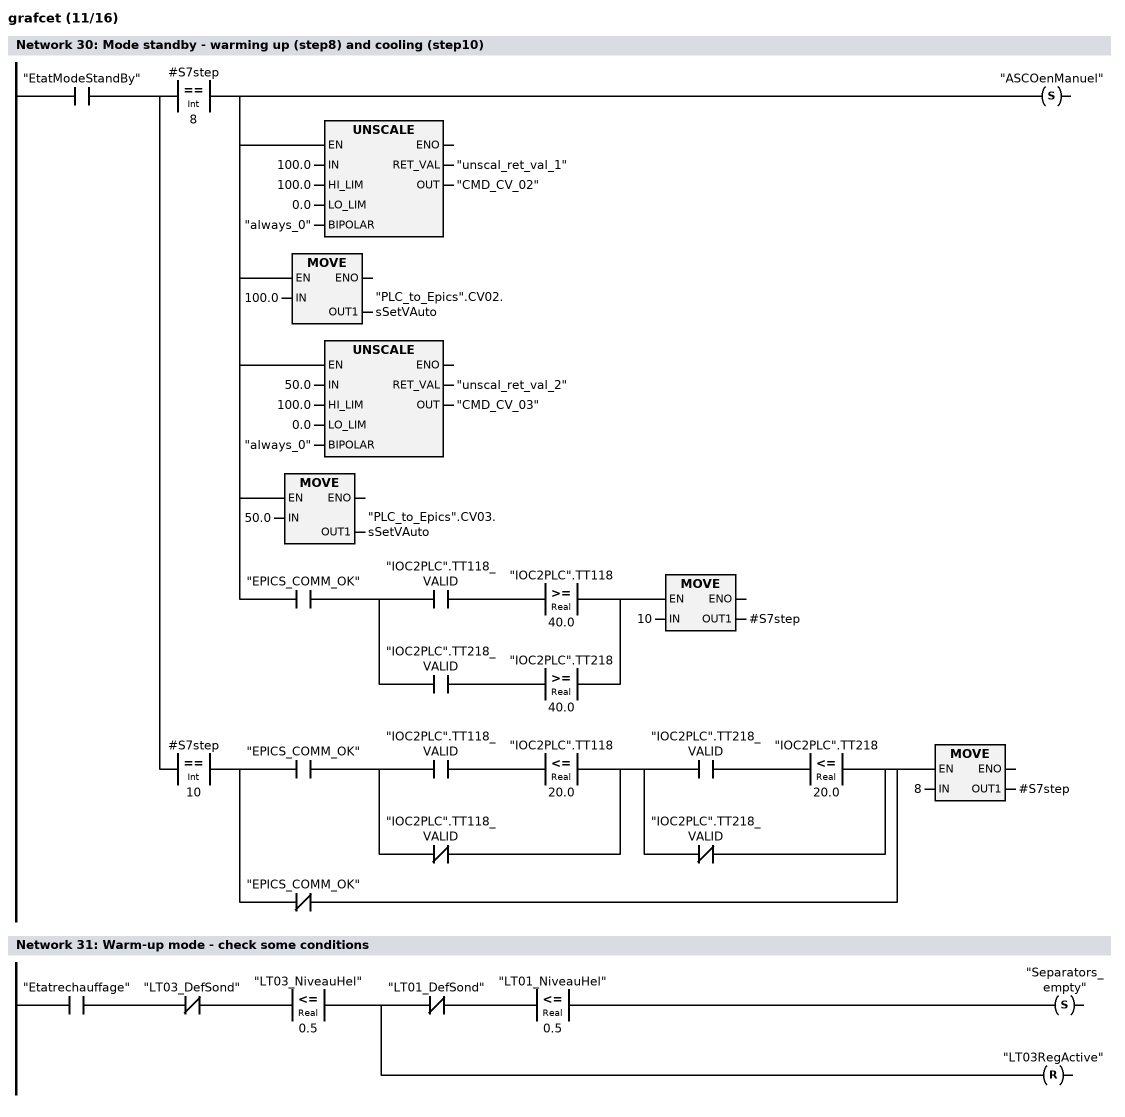
   #_w1 := "EtatModeStandBy" AND (#S7step = 8);
   IF #_w1 THEN "ASCOenManuel" := TRUE; END_IF;
   #_w2 := "EtatModeStandBy";
   IF #_w1 THEN
       "unscal_ret_val_1" := UNSCALE(IN := 100.0,
                               HI_LIM := 100.0,
                               LO_LIM := 0.0,
                               BIPOLAR := "always_0",
                               OUT => "CMD_CV_02");
       "PLC_to_Epics".CV02.sSetVAuto := 100.0;
       "unscal_ret_val_2" := UNSCALE(IN := 50.0,
                               HI_LIM := 100.0,
                               LO_LIM := 0.0,
                               BIPOLAR := "always_0",
                               OUT => "CMD_CV_03");
       "PLC_to_Epics".CV03.sSetVAuto := 50.0;
   END_IF;
   IF #_w1 AND "EPICS_COMM_OK" AND (("IOC2PLC".TT118_VALID AND ("IOC2PLC".TT118 >= 40.0)) OR ("IOC2PLC".TT218_VALID AND ("IOC2PLC".TT218 >= 40.0))) THEN
       #S7step := 10;
   END_IF;
   IF #_w2 AND (#S7step = 10) AND (("EPICS_COMM_OK" AND (("IOC2PLC".TT118_VALID AND ("IOC2PLC".TT118 <= 20.0)) OR NOT "IOC2PLC".TT118_VALID) AND (("IOC2PLC".TT218_VALID AND ("IOC2PLC".TT218 <= 20.0)) OR NOT "IOC2PLC".TT218_VALID)) OR NOT "EPICS_COMM_OK") THEN
       #S7step := 8;
   END_IF;
END_REGION

REGION Network 31: Warm-up mode - check some conditions
   #_w1 := "Etatrechauffage" AND NOT "LT03_DefSond" AND ("LT03_NiveauHel" <= 0.5);
   IF #_w1 AND NOT "LT01_DefSond" AND ("LT01_NiveauHel" <= 0.5) THEN "Separators_empty" := TRUE; END_IF;
   IF #_w1 THEN "LT03RegActive" := FALSE; END_IF;
END_REGION

REGION Network 32: Warm-up: set-up the settings of CV01-CV04
   // Set-up the settings depending on the LHe levels in the phase separators
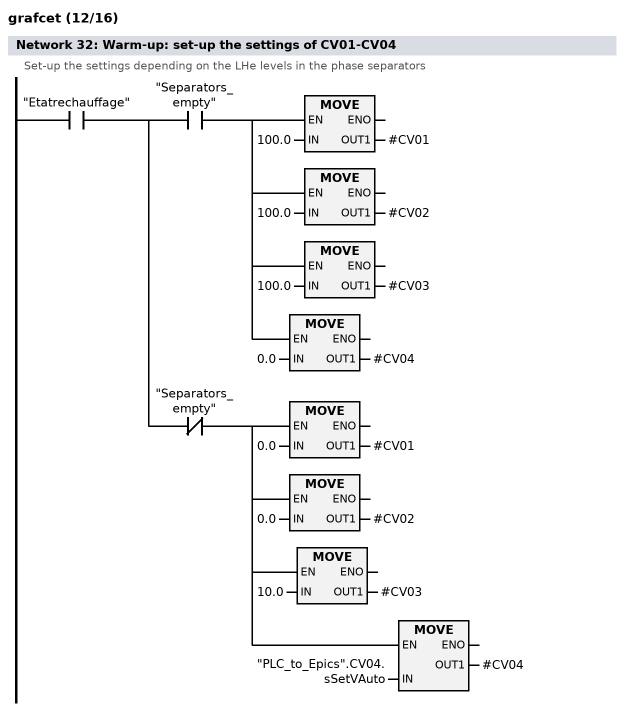
   RUNG wire#powerrail
      Contact( "Etatrechauffage" )
      wire#w1
      Contact( "Separators_empty" )
      wire#w2
      { S7_GenerateENO := "TRUE" } Move(in := 100.0, out1 => #CV01)
   END_RUNG
   RUNG wire#w2
      { S7_GenerateENO := "TRUE" } Move(in := 100.0, out1 => #CV02)
   END_RUNG
   RUNG wire#w2
      { S7_GenerateENO := "TRUE" } Move(in := 100.0, out1 => #CV03)
   END_RUNG
   RUNG wire#w2
      { S7_GenerateENO := "TRUE" } Move(in := 0.0, out1 => #CV04)
   END_RUNG
   RUNG wire#w1
      I_Contact( "Separators_empty" )
      wire#w3
      { S7_GenerateENO := "TRUE" } Move(in := 0.0, out1 => #CV01)
   END_RUNG
   RUNG wire#w3
      { S7_GenerateENO := "TRUE" } Move(in := 0.0, out1 => #CV02)
   END_RUNG
   RUNG wire#w3
      { S7_GenerateENO := "TRUE" } Move(in := 10.0, out1 => #CV03)
   END_RUNG
   RUNG wire#w3
      { S7_GenerateENO := "TRUE" } Move(in := "PLC_to_Epics".CV04.sSetVAuto, out1 => #CV04)
   END_RUNG
   // the same network as SCL:
   IF "Etatrechauffage" AND "Separators_empty" THEN
       #CV01 := 100.0;
       #CV02 := 100.0;
       #CV03 := 100.0;
       #CV04 := 0.0;
   END_IF;
   IF "Etatrechauffage" AND NOT "Separators_empty" THEN
       #CV01 := 0.0;
       #CV02 := 0.0;
       #CV03 := 10.0;
       #CV04 := "PLC_to_Epics".CV04.sSetVAuto;
   END_IF;
END_REGION

REGION Network 33: Mode Rechauffage
   // The heaters are handled in Manage_HEATERS
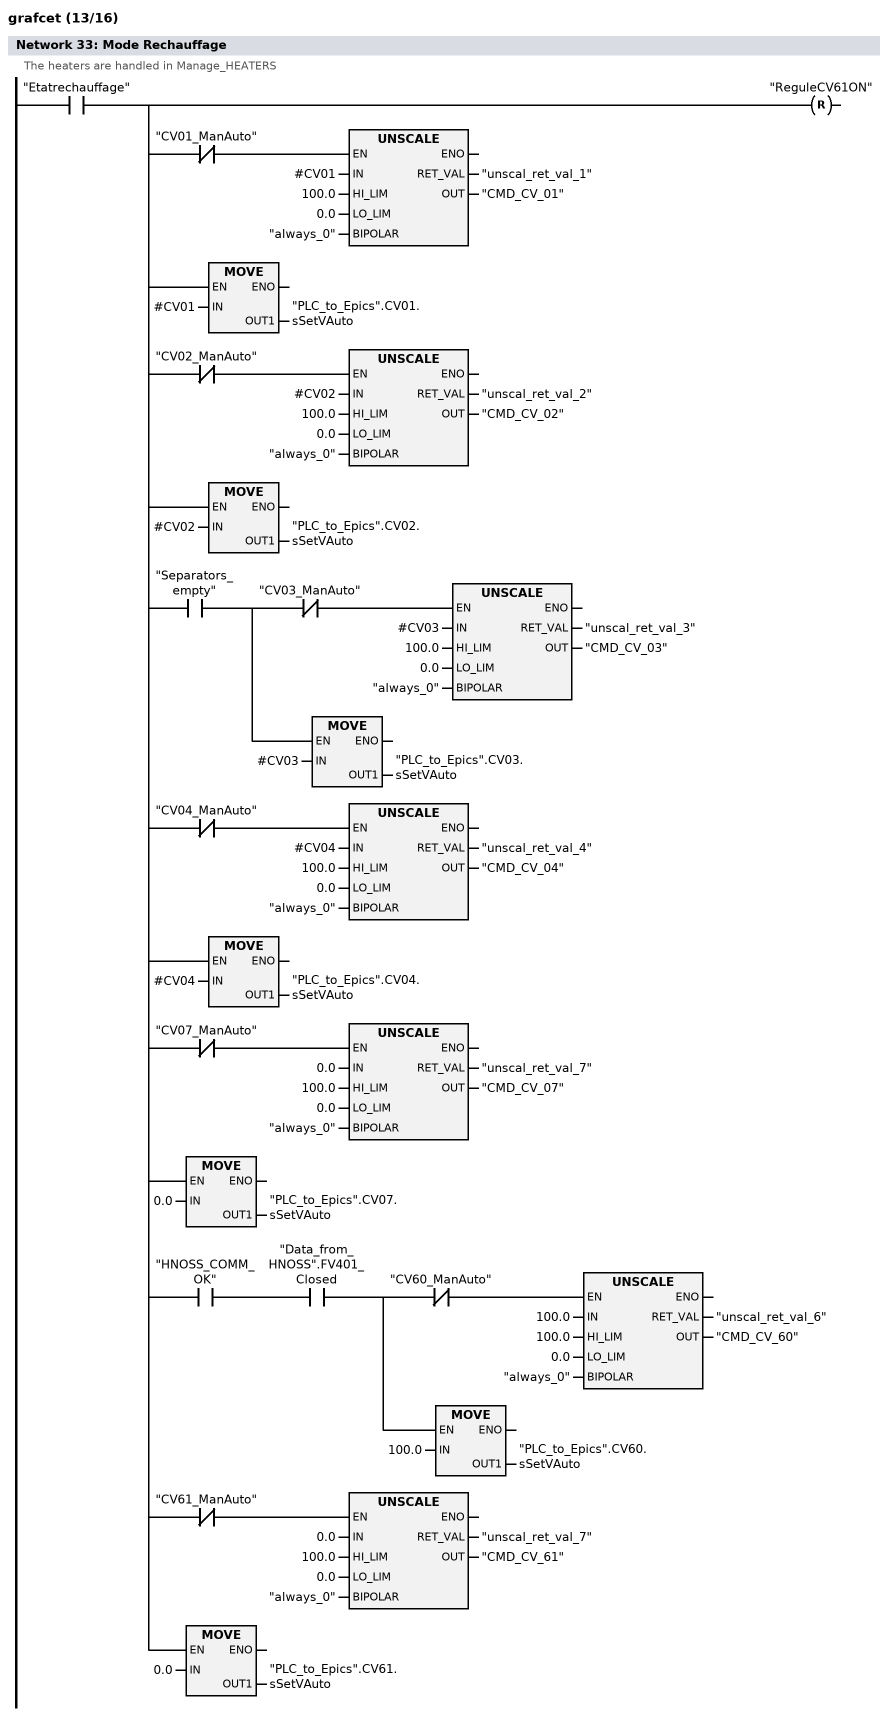
   IF "Etatrechauffage" THEN "ReguleCV61ON" := FALSE; END_IF;
   #_w1 := "Etatrechauffage";
   IF "Etatrechauffage" AND NOT "CV01_ManAuto" THEN
       "unscal_ret_val_1" := UNSCALE(IN := #CV01,
                               HI_LIM := 100.0,
                               LO_LIM := 0.0,
                               BIPOLAR := "always_0",
                               OUT => "CMD_CV_01");
   END_IF;
   IF #_w1 THEN "PLC_to_Epics".CV01.sSetVAuto := #CV01; END_IF;
   IF #_w1 AND NOT "CV02_ManAuto" THEN
       "unscal_ret_val_2" := UNSCALE(IN := #CV02,
                               HI_LIM := 100.0,
                               LO_LIM := 0.0,
                               BIPOLAR := "always_0",
                               OUT => "CMD_CV_02");
   END_IF;
   IF #_w1 THEN "PLC_to_Epics".CV02.sSetVAuto := #CV02; END_IF;
   #_w2 := #_w1 AND "Separators_empty";
   IF #_w2 AND NOT "CV03_ManAuto" THEN
       "unscal_ret_val_3" := UNSCALE(IN := #CV03,
                               HI_LIM := 100.0,
                               LO_LIM := 0.0,
                               BIPOLAR := "always_0",
                               OUT => "CMD_CV_03");
   END_IF;
   IF #_w2 THEN "PLC_to_Epics".CV03.sSetVAuto := #CV03; END_IF;
   IF #_w1 AND NOT "CV04_ManAuto" THEN
       "unscal_ret_val_4" := UNSCALE(IN := #CV04,
                               HI_LIM := 100.0,
                               LO_LIM := 0.0,
                               BIPOLAR := "always_0",
                               OUT => "CMD_CV_04");
   END_IF;
   IF #_w1 THEN "PLC_to_Epics".CV04.sSetVAuto := #CV04; END_IF;
   IF #_w1 AND NOT "CV07_ManAuto" THEN
       "unscal_ret_val_7" := UNSCALE(IN := 0.0,
                               HI_LIM := 100.0,
                               LO_LIM := 0.0,
                               BIPOLAR := "always_0",
                               OUT => "CMD_CV_07");
   END_IF;
   IF #_w1 THEN "PLC_to_Epics".CV07.sSetVAuto := 0.0; END_IF;
   #_w3 := #_w1 AND "HNOSS_COMM_OK" AND "Data_from_HNOSS".FV401_Closed;
   IF #_w3 AND NOT "CV60_ManAuto" THEN
       "unscal_ret_val_6" := UNSCALE(IN := 100.0,
                               HI_LIM := 100.0,
                               LO_LIM := 0.0,
                               BIPOLAR := "always_0",
                               OUT => "CMD_CV_60");
   END_IF;
   IF #_w3 THEN "PLC_to_Epics".CV60.sSetVAuto := 100.0; END_IF;
   IF #_w1 AND NOT "CV61_ManAuto" THEN
       "unscal_ret_val_7" := UNSCALE(IN := 0.0,
                               HI_LIM := 100.0,
                               LO_LIM := 0.0,
                               BIPOLAR := "always_0",
                               OUT => "CMD_CV_61");
   END_IF;
   IF #_w1 THEN "PLC_to_Epics".CV61.sSetVAuto := 0.0; END_IF;
END_REGION

REGION Network 34: Mode manuel ASCO
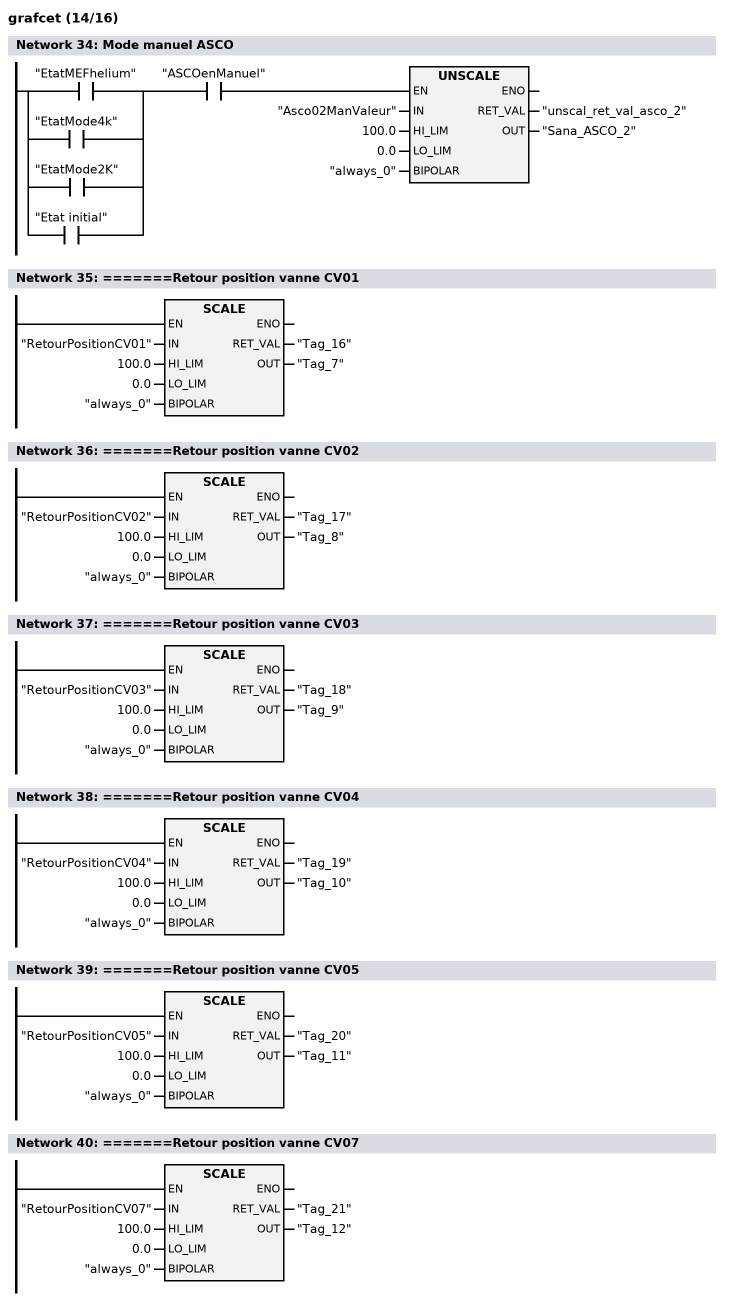
   IF ("EtatMEFhelium" OR "EtatMode4k" OR "EtatMode2K" OR "Etat initial") AND "ASCOenManuel" THEN
       "unscal_ret_val_asco_2" := UNSCALE(in := "Asco02ManValeur",
                               hi_lim := 100.0,
                               lo_lim := 0.0,
                               bipolar := "always_0",
                               out => "Sana_ASCO_2");
   END_IF;
END_REGION

REGION Network 35: =======Retour position vanne CV01
   "Tag_16" := SCALE(in := "RetourPositionCV01",
                     hi_lim := 100.0,
                     lo_lim := 0.0,
                     bipolar := "always_0",
                     out => "Tag_7");
END_REGION

REGION Network 36: =======Retour position vanne CV02
   "Tag_17" := SCALE(in := "RetourPositionCV02",
                     hi_lim := 100.0,
                     lo_lim := 0.0,
                     bipolar := "always_0",
                     out => "Tag_8");
END_REGION

REGION Network 37: =======Retour position vanne CV03
   "Tag_18" := SCALE(in := "RetourPositionCV03",
                     hi_lim := 100.0,
                     lo_lim := 0.0,
                     bipolar := "always_0",
                     out => "Tag_9");
END_REGION

REGION Network 38: =======Retour position vanne CV04
   "Tag_19" := SCALE(in := "RetourPositionCV04",
                     hi_lim := 100.0,
                     lo_lim := 0.0,
                     bipolar := "always_0",
                     out => "Tag_10");
END_REGION

REGION Network 39: =======Retour position vanne CV05
   "Tag_20" := SCALE(in := "RetourPositionCV05",
                     hi_lim := 100.0,
                     lo_lim := 0.0,
                     bipolar := "always_0",
                     out => "Tag_11");
END_REGION

REGION Network 40: =======Retour position vanne CV07
   "Tag_21" := SCALE(in := "RetourPositionCV07",
                     hi_lim := 100.0,
                     lo_lim := 0.0,
                     bipolar := "always_0",
                     out => "Tag_12");
END_REGION

REGION Network 41: =======Retour position vanne CV60
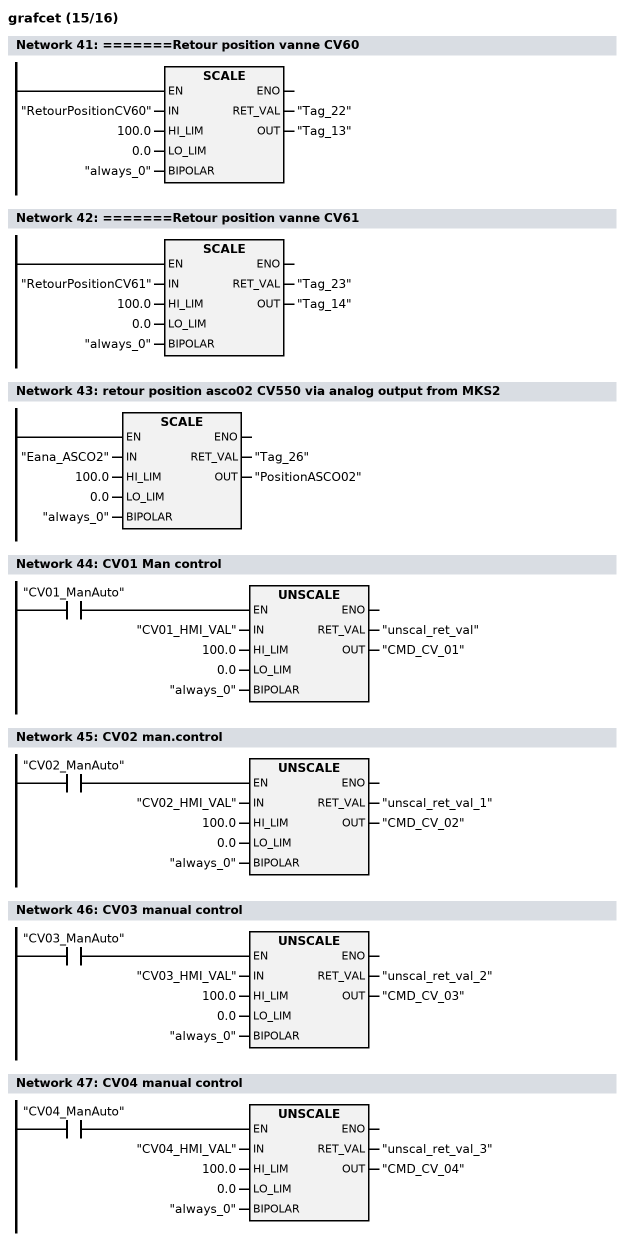
   "Tag_22" := SCALE(in := "RetourPositionCV60",
                     hi_lim := 100.0,
                     lo_lim := 0.0,
                     bipolar := "always_0",
                     out => "Tag_13");
END_REGION

REGION Network 42: =======Retour position vanne CV61
   "Tag_23" := SCALE(in := "RetourPositionCV61",
                     hi_lim := 100.0,
                     lo_lim := 0.0,
                     bipolar := "always_0",
                     out => "Tag_14");
END_REGION

REGION Network 43: retour position asco02 CV550 via analog output from MKS2
   "Tag_26" := SCALE(in := "Eana_ASCO2",
                     hi_lim := 100.0,
                     lo_lim := 0.0,
                     bipolar := "always_0",
                     out => "PositionASCO02");
END_REGION

REGION Network 44: CV01 Man control
   IF "CV01_ManAuto" THEN
       "unscal_ret_val" := UNSCALE(in := "CV01_HMI_VAL",
                               hi_lim := 100.0,
                               lo_lim := 0.0,
                               bipolar := "always_0",
                               out => "CMD_CV_01");
   END_IF;
END_REGION

REGION Network 45: CV02 man.control
   IF "CV02_ManAuto" THEN
       "unscal_ret_val_1" := UNSCALE(in := "CV02_HMI_VAL",
                               hi_lim := 100.0,
                               lo_lim := 0.0,
                               bipolar := "always_0",
                               out => "CMD_CV_02");
   END_IF;
END_REGION

REGION Network 46: CV03 manual control
   IF "CV03_ManAuto" THEN
       "unscal_ret_val_2" := UNSCALE(in := "CV03_HMI_VAL",
                               hi_lim := 100.0,
                               lo_lim := 0.0,
                               bipolar := "always_0",
                               out => "CMD_CV_03");
   END_IF;
END_REGION

REGION Network 47: CV04 manual control
   IF "CV04_ManAuto" THEN
       "unscal_ret_val_3" := UNSCALE(in := "CV04_HMI_VAL",
                               hi_lim := 100.0,
                               lo_lim := 0.0,
                               bipolar := "always_0",
                               out => "CMD_CV_04");
   END_IF;
END_REGION

REGION Network 48: CV07 manual control
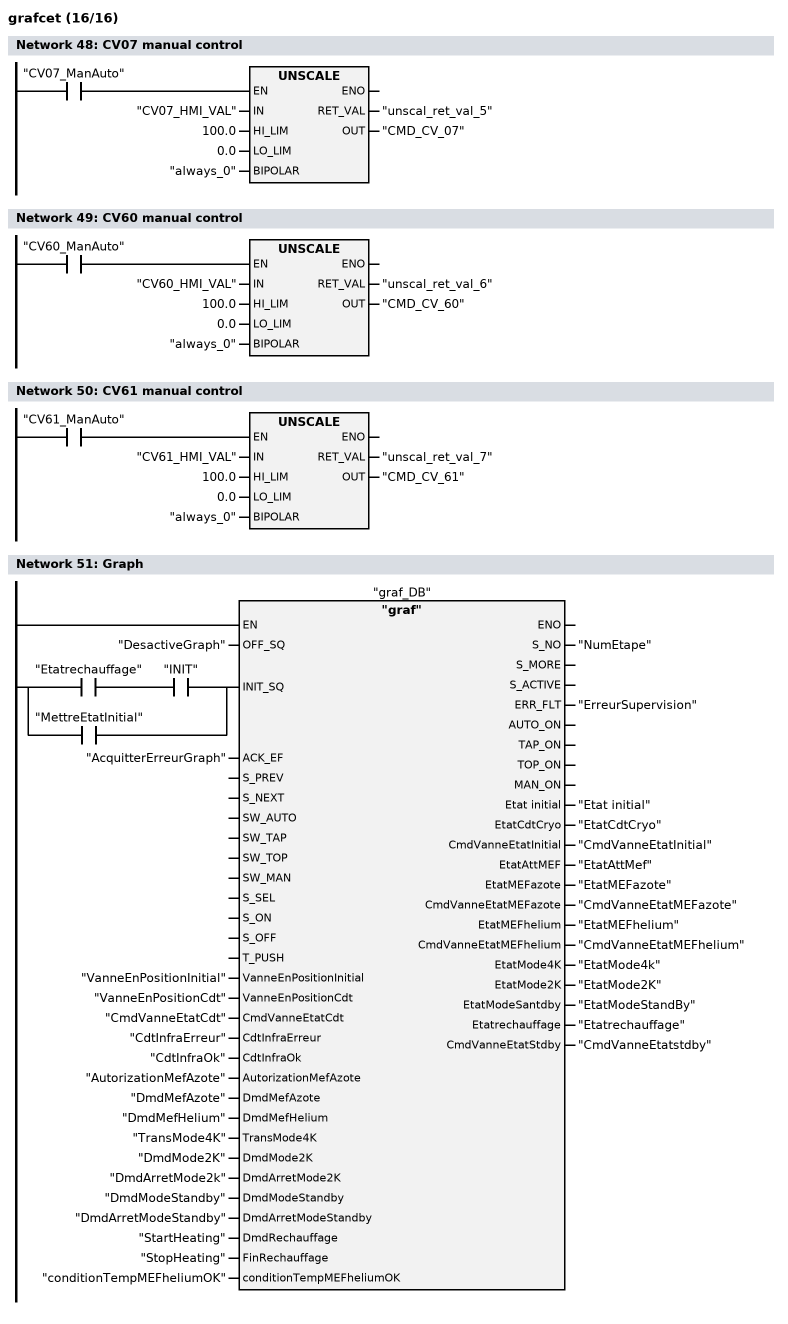
   IF "CV07_ManAuto" THEN
       "unscal_ret_val_5" := UNSCALE(in := "CV07_HMI_VAL",
                               hi_lim := 100.0,
                               lo_lim := 0.0,
                               bipolar := "always_0",
                               out => "CMD_CV_07");
   END_IF;
END_REGION

REGION Network 49: CV60 manual control
   IF "CV60_ManAuto" THEN
       "unscal_ret_val_6" := UNSCALE(in := "CV60_HMI_VAL",
                               hi_lim := 100.0,
                               lo_lim := 0.0,
                               bipolar := "always_0",
                               out => "CMD_CV_60");
   END_IF;
END_REGION

REGION Network 50: CV61 manual control
   IF "CV61_ManAuto" THEN
       "unscal_ret_val_7" := UNSCALE(in := "CV61_HMI_VAL",
                               hi_lim := 100.0,
                               lo_lim := 0.0,
                               bipolar := "always_0",
                               out => "CMD_CV_61");
   END_IF;
END_REGION

REGION Network 51: Graph
   "graf_DB"(OFF_SQ := "DesactiveGraph",   // "graf"
             INIT_SQ := "MettreEtatInitial" OR ("Etatrechauffage" AND "INIT"),
             ACK_EF := "AcquitterErreurGraph",
             VanneEnPositionInitial := "VanneEnPositionInitial",
             VanneEnPositionCdt := "VanneEnPositionCdt",
             CmdVanneEtatCdt := "CmdVanneEtatCdt",
             CdtInfraErreur := "CdtInfraErreur",
             CdtInfraOk := "CdtInfraOk",
             AutorizationMefAzote := "AutorizationMefAzote",
             DmdMefAzote := "DmdMefAzote",
             DmdMefHelium := "DmdMefHelium",
             TransMode4K := "TransMode4K",
             DmdMode2K := "DmdMode2K",
             DmdArretMode2K := "DmdArretMode2k",
             DmdModeStandby := "DmdModeStandby",
             DmdArretModeStandby := "DmdArretModeStandby",
             DmdRechauffage := "StartHeating",
             FinRechauffage := "StopHeating",
             conditionTempMEFheliumOK := "conditionTempMEFheliumOK",
             S_NO => "NumEtape",
             ERR_FLT => "ErreurSupervision",
             "Etat initial" => "Etat initial",
             EtatCdtCryo => "EtatCdtCryo",
             CmdVanneEtatInitial => "CmdVanneEtatInitial",
             EtatAttMEF => "EtatAttMef",
             EtatMEFazote => "EtatMEFazote",
             CmdVanneEtatMEFazote => "CmdVanneEtatMEFazote",
             EtatMEFhelium => "EtatMEFhelium",
             CmdVanneEtatMEFhelium => "CmdVanneEtatMEFhelium",
             EtatMode4K => "EtatMode4k",
             EtatMode2K => "EtatMode2K",
             EtatModeSantdby => "EtatModeStandBy",
             Etatrechauffage => "Etatrechauffage",
             CmdVanneEtatStdby => "CmdVanneEtatstdby");
END_REGION

REGION Network 52 (STL): Copy step numbe to HNOSS
         L     #S4step;
         T     "Data_fo_HNOSS".S4step;
         L     #S5step;
         T     "Data_fo_HNOSS".S5step;
         L     #S6step;
         T     "Data_fo_HNOSS".S6step;
         L     #S7step;
         T     "Data_fo_HNOSS".S7step;
         L     #S8step;
         T     "Data_fo_HNOSS".S8step;
         L     #S9step;
         T     "Data_fo_HNOSS".S9step;
         L     #S10step;
         T     "Data_fo_HNOSS".S10step;
         L     #Sxstep;
         T     "Data_fo_HNOSS".SXstep;
END_REGION
END_FUNCTION

FUNCTION "UpdateData2HNOSS" : Void   // FC303, LAD
{ S7_Optimized_Access := 'FALSE' }
AUTHOR : KG
VERSION : 0.1
BEGIN

REGION Network 1: Initial state
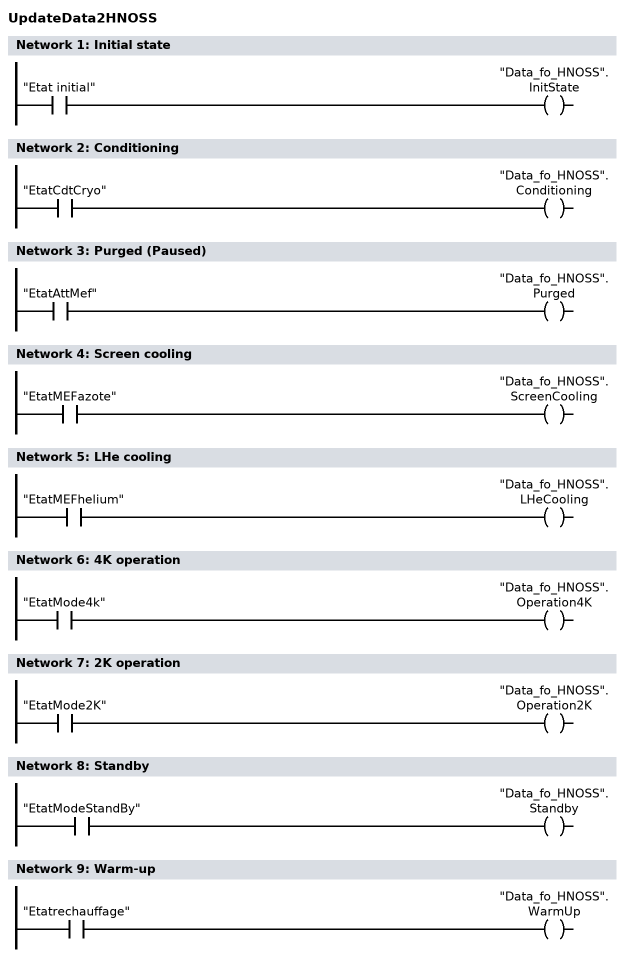
   RUNG wire#powerrail
      Contact( "Etat initial" )
      Coil( "Data_fo_HNOSS".InitState )
   END_RUNG
   // the same network as SCL:
   "Data_fo_HNOSS".InitState := "Etat initial";
END_REGION

REGION Network 2: Conditioning
   RUNG wire#powerrail
      Contact( "EtatCdtCryo" )
      Coil( "Data_fo_HNOSS".Conditioning )
   END_RUNG
   // the same network as SCL:
   "Data_fo_HNOSS".Conditioning := "EtatCdtCryo";
END_REGION

REGION Network 3: Purged (Paused)
   RUNG wire#powerrail
      Contact( "EtatAttMef" )
      Coil( "Data_fo_HNOSS".Purged )
   END_RUNG
   // the same network as SCL:
   "Data_fo_HNOSS".Purged := "EtatAttMef";
END_REGION

REGION Network 4: Screen cooling
   RUNG wire#powerrail
      Contact( "EtatMEFazote" )
      Coil( "Data_fo_HNOSS".ScreenCooling )
   END_RUNG
   // the same network as SCL:
   "Data_fo_HNOSS".ScreenCooling := "EtatMEFazote";
END_REGION

REGION Network 5: LHe cooling
   RUNG wire#powerrail
      Contact( "EtatMEFhelium" )
      Coil( "Data_fo_HNOSS".LHeCooling )
   END_RUNG
   // the same network as SCL:
   "Data_fo_HNOSS".LHeCooling := "EtatMEFhelium";
END_REGION

REGION Network 6: 4K operation
   RUNG wire#powerrail
      Contact( "EtatMode4k" )
      Coil( "Data_fo_HNOSS".Operation4K )
   END_RUNG
   // the same network as SCL:
   "Data_fo_HNOSS".Operation4K := "EtatMode4k";
END_REGION

REGION Network 7: 2K operation
   RUNG wire#powerrail
      Contact( "EtatMode2K" )
      Coil( "Data_fo_HNOSS".Operation2K )
   END_RUNG
   // the same network as SCL:
   "Data_fo_HNOSS".Operation2K := "EtatMode2K";
END_REGION

REGION Network 8: Standby
   RUNG wire#powerrail
      Contact( "EtatModeStandBy" )
      Coil( "Data_fo_HNOSS".Standby )
   END_RUNG
   // the same network as SCL:
   "Data_fo_HNOSS".Standby := "EtatModeStandBy";
END_REGION

REGION Network 9: Warm-up
   RUNG wire#powerrail
      Contact( "Etatrechauffage" )
      Coil( "Data_fo_HNOSS".WarmUp )
   END_RUNG
   // the same network as SCL:
   "Data_fo_HNOSS".WarmUp := "Etatrechauffage";
END_REGION
END_FUNCTION

FUNCTION "#FC_CONTROL_HEATER" : Void   // FC313, STL
TITLE = Object : Heater
{ S7_Optimized_Access := 'FALSE' }
VERSION : 0.1
BEGIN

REGION Network 1: Initialise of Equipment
         A     "INIT";
         JCN   INIT;
         S     #Object.XH;
   INIT: NOP   0;
END_REGION

REGION Network 2: Epics Commands
   //Set Auto
         A     #cmdEpics.cmdAuto;
         S     #Object.XH;

   // Set Manu
         A     #cmdEpics.cmdMan;
         R     #Object.XH;

   // Set manual command
         A     #cmdEpics.cmdSet;
         S     #Object.H;

   // Reset manual command
         A     #cmdEpics.cmdRst;
         R     #Object.H;

   // Set High limit
         A     #cmdEpics.cmdHL;
         JCN   Epc0;
         L     #cmdEpics.cHL;
         T     #Object.Tt_Max;
   Epc0: NOP   0;

   // Set Low limit
         A     #cmdEpics.cmdLL;
         JCN   Epc1;
         L     #cmdEpics.cLL;
         T     #Object.Tt_Min;
   Epc1: NOP   0;

   EP01: NOP   0;

   // Reset Epics Commands
         R     #cmdEpics.cmdAuto;
         R     #cmdEpics.cmdMan;
         R     #cmdEpics.cmdSet;
         R     #cmdEpics.cmdRst;
         R     #cmdEpics.cmdHL;
         R     #cmdEpics.cmdLL;
END_REGION

REGION Network 3: Data acquisition
   //Input Temperature
         L     #TtA;
         T     #Object.ValueA;

         L     #TtB;
         T     #Object.ValueB;

         L     #TtC;
         T     #Object.ValueC;

         L     #TtD;
         T     #Object.ValueD;

         L     #TtE;
         T     #Object.ValueE;

         L     #TtF;
         T     #Object.ValueF;


   // Termoswitch
         AN    #TS;
         =     #Object.TS;

   // External Command
         A     #ExtCmd;
         =     #Object.R_ExtCmd;

   //Number of Temperature
         L     #Nb_Tt;
         T     #Object.Nb_Tt;
END_REGION

REGION Network 4: Management Thermoswitch
   //ThermoSwitch
   //Timer On
         A     #Object.TS;
         =     #Rec_Ts_On;

         CALL  "#FC_TIMER"
         ( Input     := #Rec_Ts_On,
           Input_RTZ := FALSE,
           Pulse     := "oneSecPls",
           RTZ       := FALSE,
           Tbase     := 1,
           Preset1   := #Object.P_TS_Ton,
           Preset2   := #T_Time,
           Time1     := #Object.TS_Ton,
           Time2     := #T_Time
         );

         L     #Object.TS_Ton;
         L     #Object.P_TS_Ton;
         >=D;
         S     #Object.TS_Calc;

   //Timer Off
         AN    #Object.TS;
         =     #Rec_Ts_Off;

         CALL  "#FC_TIMER"
         ( Input     := #Rec_Ts_Off,
           Input_RTZ := FALSE,
           Pulse     := "oneSecPls",
           RTZ       := FALSE,
           Tbase     := 1,
           Preset1   := #Object.P_TS_Toff,
           Preset2   := #T_Time,
           Time1     := #Object.TS_Toff,
           Time2     := #T_Time
         );

         L     #Object.TS_Toff;
         L     #Object.P_TS_Toff;
         >=D;
         R     #Object.TS_Calc;
END_REGION

REGION Network 5: Equipment Pilot Command
   //Test of number of temperature to SET
         A(;
         L     #Nb_Tt;
         L     1;
         ==I;
         );
         JC    T01S;
         A(;
         L     #Nb_Tt;
         L     2;
         ==I;
         );
         JC    T02S;
         A(;
         L     #Nb_Tt;
         L     3;
         ==I;
         );
         JC    T03S;
         A(;
         L     #Nb_Tt;
         L     4;
         ==I;
         );
         JC    T04S;
         A(;
         L     #Nb_Tt;
         L     5;
         ==I;
         );
         JC    T05S;
         A(;
         L     #Nb_Tt;
         L     6;
         ==I;
         );
         JC    T06S;

         JU    NCS;

   //Set Command
   T06S: A(;
         L     #Object.ValueF;
         L     #Object.Tt_Min;
         <R;
         );
         S     #Object.Pilot;

   T05S: A(;
         L     #Object.ValueE;
         L     #Object.Tt_Min;
         <R;
         );
         S     #Object.Pilot;

   T04S: A(;
         L     #Object.ValueD;
         L     #Object.Tt_Min;
         <R;
         );
         S     #Object.Pilot;

   T03S: A(;
         L     #Object.ValueC;
         L     #Object.Tt_Min;
         <R;
         );
         S     #Object.Pilot;

   T02S: A(;
         L     #Object.ValueB;
         L     #Object.Tt_Min;
         <R;
         );
         S     #Object.Pilot;

   T01S: A(;
         L     #Object.ValueA;
         L     #Object.Tt_Min;
         <R;
         );
         S     #Object.Pilot;

   NCS:  NOP   0;


   //Test of number of temperature to RESET
         A(;
         L     #Nb_Tt;
         L     1;
         ==I;
         );
         JC    T01R;
         A(;
         L     #Nb_Tt;
         L     2;
         ==I;
         );
         JC    T02R;
         A(;
         L     #Nb_Tt;
         L     3;
         ==I;
         );
         JC    T03R;
         A(;
         L     #Nb_Tt;
         L     4;
         ==I;
         );
         JC    T04R;
         A(;
         L     #Nb_Tt;
         L     5;
         ==I;
         );
         JC    T05R;
         A(;
         L     #Nb_Tt;
         L     6;
         ==I;
         );
         JC    T06R;


   //Reset Command
   T06R: A(;
         L     #Object.ValueF;
         L     #Object.Tt_Max;
         >=R;
         );
         R     #Object.Pilot;

   T05R: A(;
         L     #Object.ValueE;
         L     #Object.Tt_Max;
         >=R;
         );
         R     #Object.Pilot;

   T04R: A(;
         L     #Object.ValueD;
         L     #Object.Tt_Max;
         >=R;
         );
         R     #Object.Pilot;

   T03R: A(;
         L     #Object.ValueC;
         L     #Object.Tt_Max;
         >=R;
         );
         R     #Object.Pilot;

   T02R: A(;
         L     #Object.ValueB;
         L     #Object.Tt_Max;
         >=R;
         );
         R     #Object.Pilot;

   T01R: A(;
         L     #Object.ValueA;
         L     #Object.Tt_Max;
         >=R;
         );
         R     #Object.Pilot;
END_REGION

REGION Network 6: External Pilot
   // External Forcage command
         A     #Object.R_ExtCmd;
         JCN   ExtF;
         S     #Object.Pilot;
   ExtF: NOP   0;
END_REGION

REGION Network 7: Delay of Command
   //Timer On
         A(;
         A     #Object.XH;
         A     #Object.X;
         O;
         AN    #Object.XH;
         A     #Object.H;
         );
         AN    #Object.TS_Calc;
         A     #Object.Pilot;
         =     #Rec_Pilot_On;

         CALL  "#FC_TIMER"
         ( Input     := #Rec_Pilot_On,
           Input_RTZ := FALSE,
           Pulse     := "oneSecPls",
           RTZ       := FALSE,
           Tbase     := 1,
           Preset1   := #Object.P_Pilot_Ton,
           Preset2   := #T_Time,
           Time1     := #Object.Pilot_Ton,
           Time2     := #T_Time
         );

         A(;
         L     #Object.Pilot_Ton;
         L     #Object.P_Pilot_Ton;
         >=D;
         );
         =     #Object.Pilot_Calc;

   // Output command
         A     #Object.Pilot_Calc;
         =     #EH;
         =     #Object.R_EH;
END_REGION

REGION Network 8: Auto copy command on the hand control
         A     #Object.XH;
         A     #Object.R_EH;
         S     #Object.H;

         A     #Object.XH;
         AN    #Object.R_EH;
         R     #Object.H;
END_REGION

REGION Network 9: Equipement ok
         A     #Object.XH;
         =     #Object.Ok;
END_REGION

REGION Network 10: Temps d'utilisation
         CALL  "#FC_TIMER"
         ( Input     := #Object.R_EH,
           Input_RTZ := #Object.Raz_Fct_Run,
           Pulse     := "oneSecPls",
           RTZ       := TRUE,
           Tbase     := 1,
           Preset1   := 2073600000,
           Preset2   := #T_Time,
           Time1     := #Object.T_run,
           Time2     := #T_Time
         );
END_REGION

REGION Network 11: Epics State
   // Copy of Auto/Manual mode
         A     #Object.XH;
         =     #sEpics.sAuto;

   // Copy of ThermoSwitch
         A     #Object.TS;
         =     #sEpics.sTsw;

   // Copy of Heater On signal
         A     #Object.R_EH;
         =     #sEpics.sHtrOn;

   // Copy of Command in Auto Mode
         A     #Object.X;
         =     #sEpics.sCmdAuto;

   // Copy of Command
         A(;
         A     #Object.XH;
         A     #Object.X;
         O;
         AN    #Object.XH;
         A     #Object.H;
         );
         =     #sEpics.sCmd;

   // Copy of High Limit
         L     #Object.Tt_Max;
         T     #sEpics.sHL;

   // Copy of Low Limit
         L     #Object.Tt_Min;
         T     #sEpics.sLL;
END_REGION

REGION Network 12: Reset action bool
         SET;
         R     #Object.Raz_Fct_Run;
END_REGION
END_FUNCTION

FUNCTION "#FC_TIMER" : Void   // FC323, LAD
TITLE = Object : Timer
{ S7_Optimized_Access := 'FALSE' }
AUTHOR : ISIITECH
VERSION : 0.1
// ISIITECH - Timer
// 19.01.2010 version 1.0
BEGIN

REGION Network 1 (STL): T
         A     #Input;
         JCN   ST1;
         L     #Time1;
         L     #Preset1;
         <D;
         JCN   ST2;
         A     #Pulse;
         JCN   ST2;
         L     #Time1;
         L     #Tbase;
         +D;
         T     #Time1;
         JU    ST2;
   ST1:  NOP   0;
   ST2:  NOP   0;



         A(;
         A     #RTZ;
         A     #Input_RTZ;
         );
         O(;
         AN    #Input;
         AN    #RTZ;
         );
         JCN   ST3;
         L     0;
         T     #Time1;
   ST3:  NOP   0;
END_REGION

REGION Network 2 (STL): T
         A     #Input;
         JCN   ST21;
         L     #Time2;
         L     #Preset2;
         <D;
         JCN   ST22;
         A     "point1secPls";
         JCN   ST22;
         L     #Time2;
         L     DINT#100;
         +D;
         T     #Time2;
         JU    ST22;
   ST21: NOP   0;
   ST22: NOP   0;



         A(;
         A     #RTZ;
         A     #Input_RTZ;
         );
         O(;
         AN    #Input;
         AN    #RTZ;
         );
         JCN   ST23;
         L     0;
         T     #Time2;
   ST23: NOP   0;
END_REGION
END_FUNCTION

FUNCTION "INST_CONTROL_HEATER" : Void   // FC413, LAD
TITLE = Heater controllers
{ S7_Optimized_Access := 'FALSE' }
AUTHOR : KG
VERSION : 0.1
BEGIN

REGION Network 1 (STL): Init variables
   // Dewar, Electrical Heater
         L     500.0;
         T     #Unused_TT;
         R     #ExtCmd;
END_REGION

REGION Network 2 (STL): EH90 - VB channel 1
   // Dewar, Electrical Heater
         L     2;
         T     "#DATA_HEATERS".EH90.P_TS_Ton;
         T     "#DATA_HEATERS".EH90.P_Pilot_Ton;
         L     5;
         T     "#DATA_HEATERS".EH90.P_TS_Toff;

         SET;
         A     "IOC2PLC".TT900_VALID;
         A     "EPICS_COMM_OK";
         =     #TS;

   // Force the heater ON when the temperature data is not valid
   // (TS = FALSE). The heater will be turned on for 30 s and TS
   // will be forced TRUE for 30 s. This will hopefully raise the
   // temperature enough for Pt100 to be in range (>73 K)
         SET;
         AN    #TS;
         A(;
         A     "#DATA_HEATERS".EH90.XH;
         A     "#DATA_HEATERS".EH90.X;
         O;
         AN    "#DATA_HEATERS".EH90.XH;
         A     "#DATA_HEATERS".EH90.H;
         );
         =     #ExtCmdTrig;
         CALL  TP, "IEC_Timer_EH90_DB"
         ( IN := #ExtCmdTrig,
           PT := T#30s,
           Q  := #ExtCmd,
           ET := #tmp_et
         );
         A     #ExtCmd;
         S     #TS;

         CALL  "#FC_CONTROL_HEATER"
         ( TtA      := "IOC2PLC".TT900,
           TtB      := #Unused_TT,
           TtC      := #Unused_TT,
           TtD      := #Unused_TT,
           TtE      := #Unused_TT,
           TtF      := #Unused_TT,
           Nb_Tt    := 1,
           TS       := #TS,
           ExtCmd   := #ExtCmd,
           cmdEpics := "Epics_to_PLC".EH90,
           EH       := "voie 1 chaufferette BV",
           sEpics   := "PLC_to_Epics".EH90,
           Object   := "#DATA_HEATERS".EH90
         );
END_REGION

REGION Network 3 (STL): EH93-96 - VB channel 2
   // Dewar, Electrical Heater
         L     2;
         T     "#DATA_HEATERS"."EH93-96".P_TS_Ton;
         T     "#DATA_HEATERS"."EH93-96".P_Pilot_Ton;
         L     5;
         T     "#DATA_HEATERS"."EH93-96".P_TS_Toff;

         SET;
         A     "IOC2PLC".TT930_VALID;
         A     "IOC2PLC".TT940_VALID;
         A     "IOC2PLC".TT950_VALID;
         A     "IOC2PLC".TT960_VALID;
         A     "EPICS_COMM_OK";
         =     #TS;

   // Force the heater ON when the temperature data is not valid
   // (TS = FALSE). The heater will be turned on for 30 s and TS
   // will be forced TRUE for 30 s. This will hopefully raise the
   // temperature enough for Pt100 to be in range (>73 K)
         SET;
         AN    #TS;
         A(;
         A     "#DATA_HEATERS"."EH93-96".XH;
         A     "#DATA_HEATERS"."EH93-96".X;
         O;
         AN    "#DATA_HEATERS"."EH93-96".XH;
         A     "#DATA_HEATERS"."EH93-96".H;
         );
         =     #ExtCmdTrig;
         CALL  TP , "IEC_Timer_EH93-96_DB"
         ( IN := #ExtCmdTrig,
           PT := T#30s,
           Q  := #ExtCmd,
           ET := #tmp_et
         );
         A     #ExtCmd;
         S     #TS;

         CALL  "#FC_CONTROL_HEATER"
         ( TtA      := "IOC2PLC".TT930,
           TtB      := "IOC2PLC".TT940,
           TtC      := "IOC2PLC".TT950,
           TtD      := "IOC2PLC".TT960,
           TtE      := #Unused_TT,
           TtF      := #Unused_TT,
           Nb_Tt    := 4,
           TS       := #TS,
           ExtCmd   := #ExtCmd,
           cmdEpics := "Epics_to_PLC"."EH93-96",
           EH       := "voie 2 chaufferette BV",
           sEpics   := "PLC_to_Epics"."EH93-96",
           Object   := "#DATA_HEATERS"."EH93-96"
         );
END_REGION

REGION Network 4 (STL): EH63_64_70 - VB channel 3
   // Dewar, Electrical Heater
         L     2;
         T     "#DATA_HEATERS"."EH63-70".P_TS_Ton;


         T     "#DATA_HEATERS"."EH63-70".P_Pilot_Ton;
         L     5;
         T     "#DATA_HEATERS"."EH63-70".P_TS_Toff;

         SET;
         A     "IOC2PLC".TT630_VALID;
         A     "IOC2PLC".TT640_VALID;
         A     "IOC2PLC".TT700_VALID;
         A     "EPICS_COMM_OK";
         =     #TS;
   // Force the heater ON when the temperature data is not valid
   // (TS = FALSE). The heater will be turned on for 30 s and TS
   // will be forced TRUE for 30 s. This will hopefully raise the
   // temperature enough for Pt100 to be in range (>73 K)
         SET;
         AN    #TS;
         A(;
         A     "#DATA_HEATERS"."EH63-70".XH;
         A     "#DATA_HEATERS"."EH63-70".X;
         O;
         AN    "#DATA_HEATERS"."EH63-70".XH;
         A     "#DATA_HEATERS"."EH63-70".H;
         );
         =     #ExtCmdTrig;
         CALL  TP , "IEC_Timer_EH63-70_DB"
         ( IN := #ExtCmdTrig,
           PT := T#30s,
           Q  := #ExtCmd,
           ET := #tmp_et
         );
         A     #ExtCmd;
         S     #TS;

         CALL  "#FC_CONTROL_HEATER"
         ( TtA      := "IOC2PLC".TT630,
           TtB      := "IOC2PLC".TT640,
           TtC      := "IOC2PLC".TT700,
           TtD      := #Unused_TT,
           TtE      := #Unused_TT,
           TtF      := #Unused_TT,
           Nb_Tt    := 3,
           TS       := #TS,
           ExtCmd   := #ExtCmd,
           cmdEpics := "Epics_to_PLC"."EH63-70",
           EH       := "voie 3 chaufferette BV",
           sEpics   := "PLC_to_Epics"."EH63-70",
           Object   := "#DATA_HEATERS"."EH63-70"
         );
END_REGION

REGION Network 5 (STL): EH61-62 - VB channel 4
   // Dewar, Electrical Heater
         L     2;
         T     "#DATA_HEATERS"."EH61-62".P_TS_Ton;